REGION Network 10
   RUNG wire#powerrail
      { S7_Templates := "SrcType := Real"; S7_GenerateENO := "TRUE" } Sub(in1 := "DB122".Static_0, in2 := "DB122".Static_24, out => "DB122".Static_18)
      wire#w1
      Coil( "Tag_6" )
   END_RUNG
   RUNG wire#powerrail
      { S7_Templates := "SrcType := Real"; S7_GenerateENO := "TRUE" } Sub(in1 := "DB122".Static_1, in2 := "DB122".Static_24, out => "DB122".Static_19)
   END_RUNG wire#w1
   RUNG wire#powerrail
      { S7_Templates := "SrcType := Real"; S7_GenerateENO := "TRUE" } Sub(in1 := "DB122".Static_2, in2 := "DB122".Static_24, out => "DB122".Static_20)
   END_RUNG wire#w1
   RUNG wire#powerrail
      { S7_Templates := "SrcType := Real"; S7_GenerateENO := "TRUE" } Sub(in1 := "DB122".Static_3, in2 := "DB122".Static_24, out => "DB122".Static_21)
   END_RUNG wire#w1
   RUNG wire#powerrail
      { S7_Templates := "SrcType := Real"; S7_GenerateENO := "TRUE" } Sub(in1 := "DB122".Static_4, in2 := "DB122".Static_24, out => "DB122".Static_22)
   END_RUNG wire#w1
   RUNG wire#powerrail
      { S7_Templates := "SrcType := Real"; S7_GenerateENO := "TRUE" } Sub(in1 := "DB122".Static_5, in2 := "DB122".Static_24, out => "DB122".Static_23)
   END_RUNG wire#w1
   // the same network as SCL:
   // ENO of a box is taken as its EN; it also drops when the box reports an error
   "DB122".Static_18 := "DB122".Static_0 - "DB122".Static_24;
   "DB122".Static_19 := "DB122".Static_1 - "DB122".Static_24;
   "DB122".Static_20 := "DB122".Static_2 - "DB122".Static_24;
   "DB122".Static_21 := "DB122".Static_3 - "DB122".Static_24;
   "DB122".Static_22 := "DB122".Static_4 - "DB122".Static_24;
   "DB122".Static_23 := "DB122".Static_5 - "DB122".Static_24;
   "Tag_6" := TRUE OR TRUE OR TRUE OR TRUE OR TRUE OR TRUE;
END_REGION

REGION Network 11 (STL)
         A     "MC003_EV";
         A(;
         A(;
         L     "DB121".Static_62;
         L     1;
         ==R;
         );
         A(;
         L     "DB52".Static_13;
         L     "DB122".Static_18;
         >=R;
         );
         O;
         A(;
         L     "DB121".Static_62;
         L     2;
         ==R;
         );
         A(;
         L     "DB52".Static_13;
         L     "DB122".Static_19;
         >=R;
         );
         O;
         A(;
         L     "DB121".Static_62;
         L     3;
         ==R;
         );
         A(;
         L     "DB52".Static_13;
         L     "DB122".Static_20;
         >=R;
         );
         O;
         A(;
         L     "DB121".Static_62;
         L     4;
         ==R;
         );
         A(;
         L     "DB52".Static_13;
         L     "DB122".Static_21;
         >=R;
         );
         O;
         A(;
         L     "DB121".Static_62;
         L     5;
         ==R;
         );
         A(;
         L     "DB52".Static_13;
         L     "DB122".Static_22;
         >=R;
         );
         O;
         A(;
         L     "DB121".Static_62;
         L     6;
         ==R;
         );
         A(;
         L     "DB52".Static_13;
         L     "DB122".Static_23;
         >=R;
         );
         );
         L     S5T#30S;
         SF    "Tag_13";
         NOP   0;
         NOP   0;
         NOP   0;
         A     "Tag_13";
         =     #Temp_0;
END_REGION

REGION Network 12
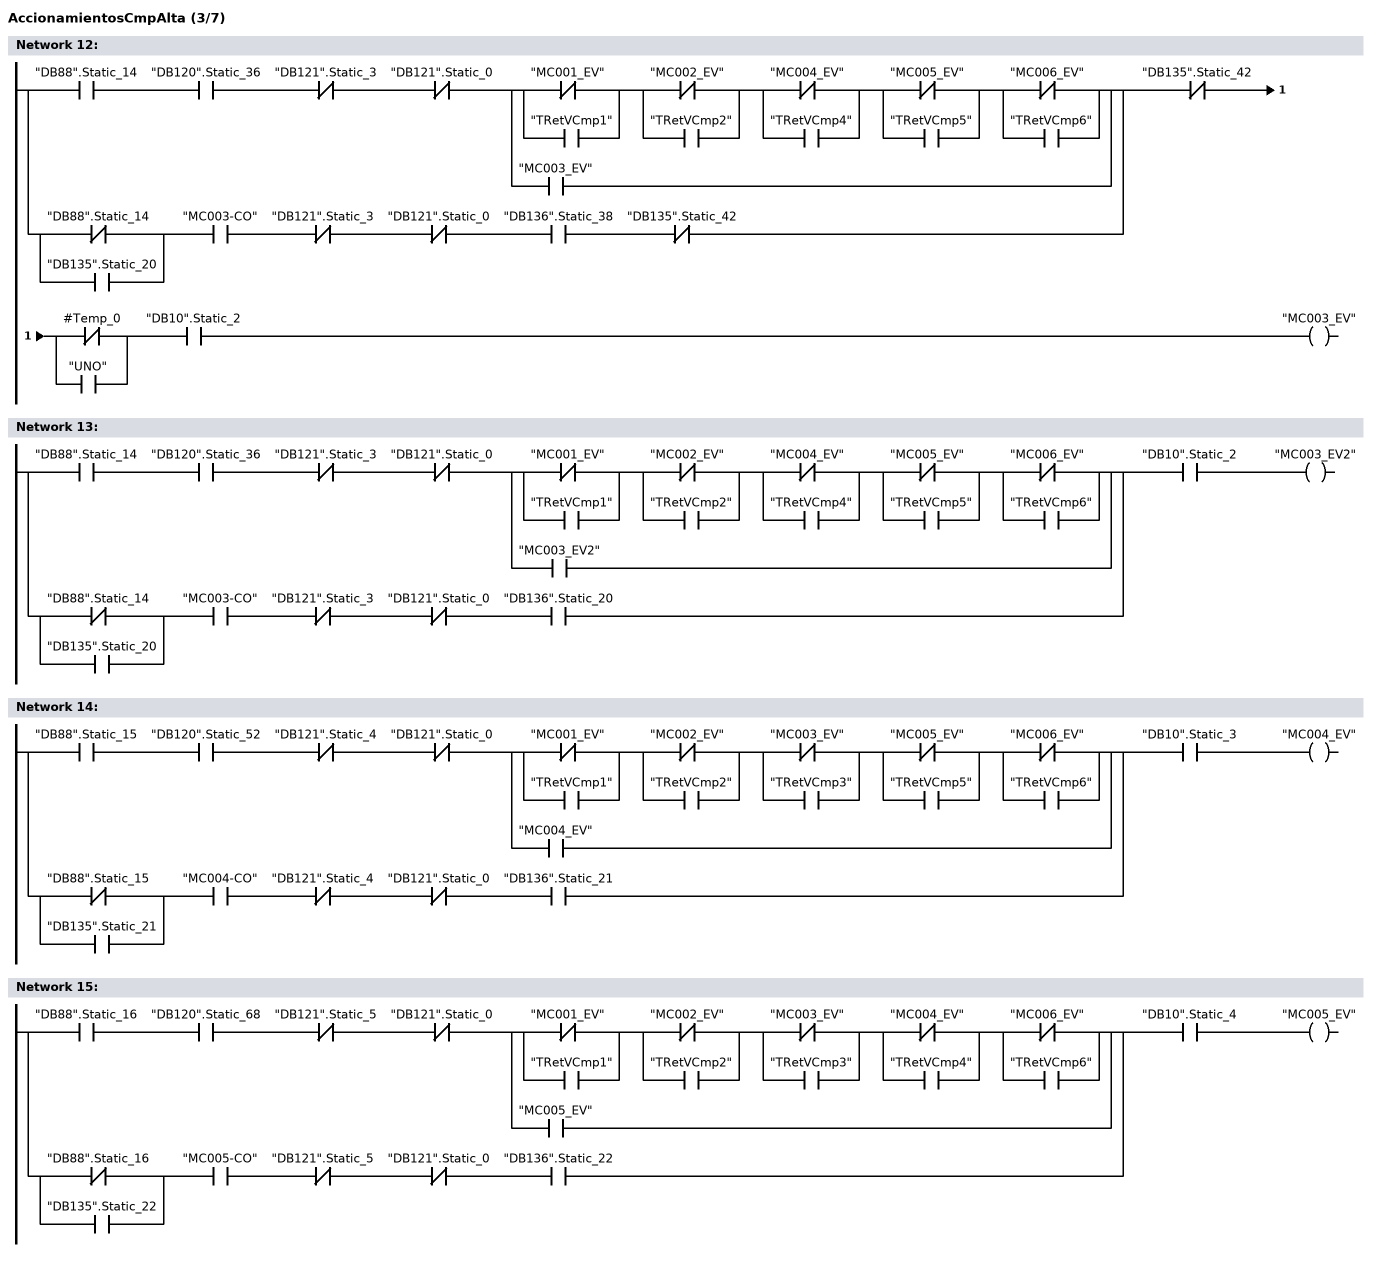
   "MC003_EV" := (("DB88".Static_14 AND "DB120".Static_36 AND NOT "DB121".Static_3 AND NOT "DB121".Static_0 AND (((NOT "MC001_EV" OR "TRetVCmp1") AND (NOT "MC002_EV" OR "TRetVCmp2") AND (NOT "MC004_EV" OR "TRetVCmp4") AND (NOT "MC005_EV" OR "TRetVCmp5") AND (NOT "MC006_EV" OR "TRetVCmp6")) OR "MC003_EV")) OR ((NOT "DB88".Static_14 OR "DB135".Static_20) AND "MC003-CO" AND NOT "DB121".Static_3 AND NOT "DB121".Static_0 AND "DB136".Static_38 AND NOT "DB135".Static_42)) AND NOT "DB135".Static_42 AND (NOT #Temp_0 OR "UNO") AND "DB10".Static_2;
END_REGION

REGION Network 13
   "MC003_EV2" := (("DB88".Static_14 AND "DB120".Static_36 AND NOT "DB121".Static_3 AND NOT "DB121".Static_0 AND (((NOT "MC001_EV" OR "TRetVCmp1") AND (NOT "MC002_EV" OR "TRetVCmp2") AND (NOT "MC004_EV" OR "TRetVCmp4") AND (NOT "MC005_EV" OR "TRetVCmp5") AND (NOT "MC006_EV" OR "TRetVCmp6")) OR "MC003_EV2")) OR ((NOT "DB88".Static_14 OR "DB135".Static_20) AND "MC003-CO" AND NOT "DB121".Static_3 AND NOT "DB121".Static_0 AND "DB136".Static_20)) AND "DB10".Static_2;
END_REGION

REGION Network 14
   "MC004_EV" := (("DB88".Static_15 AND "DB120".Static_52 AND NOT "DB121".Static_4 AND NOT "DB121".Static_0 AND (((NOT "MC001_EV" OR "TRetVCmp1") AND (NOT "MC002_EV" OR "TRetVCmp2") AND (NOT "MC003_EV" OR "TRetVCmp3") AND (NOT "MC005_EV" OR "TRetVCmp5") AND (NOT "MC006_EV" OR "TRetVCmp6")) OR "MC004_EV")) OR ((NOT "DB88".Static_15 OR "DB135".Static_21) AND "MC004-CO" AND NOT "DB121".Static_4 AND NOT "DB121".Static_0 AND "DB136".Static_21)) AND "DB10".Static_3;
END_REGION

REGION Network 15
   "MC005_EV" := (("DB88".Static_16 AND "DB120".Static_68 AND NOT "DB121".Static_5 AND NOT "DB121".Static_0 AND (((NOT "MC001_EV" OR "TRetVCmp1") AND (NOT "MC002_EV" OR "TRetVCmp2") AND (NOT "MC003_EV" OR "TRetVCmp3") AND (NOT "MC004_EV" OR "TRetVCmp4") AND (NOT "MC006_EV" OR "TRetVCmp6")) OR "MC005_EV")) OR ((NOT "DB88".Static_16 OR "DB135".Static_22) AND "MC005-CO" AND NOT "DB121".Static_5 AND NOT "DB121".Static_0 AND "DB136".Static_22)) AND "DB10".Static_4;
END_REGION

REGION Network 16
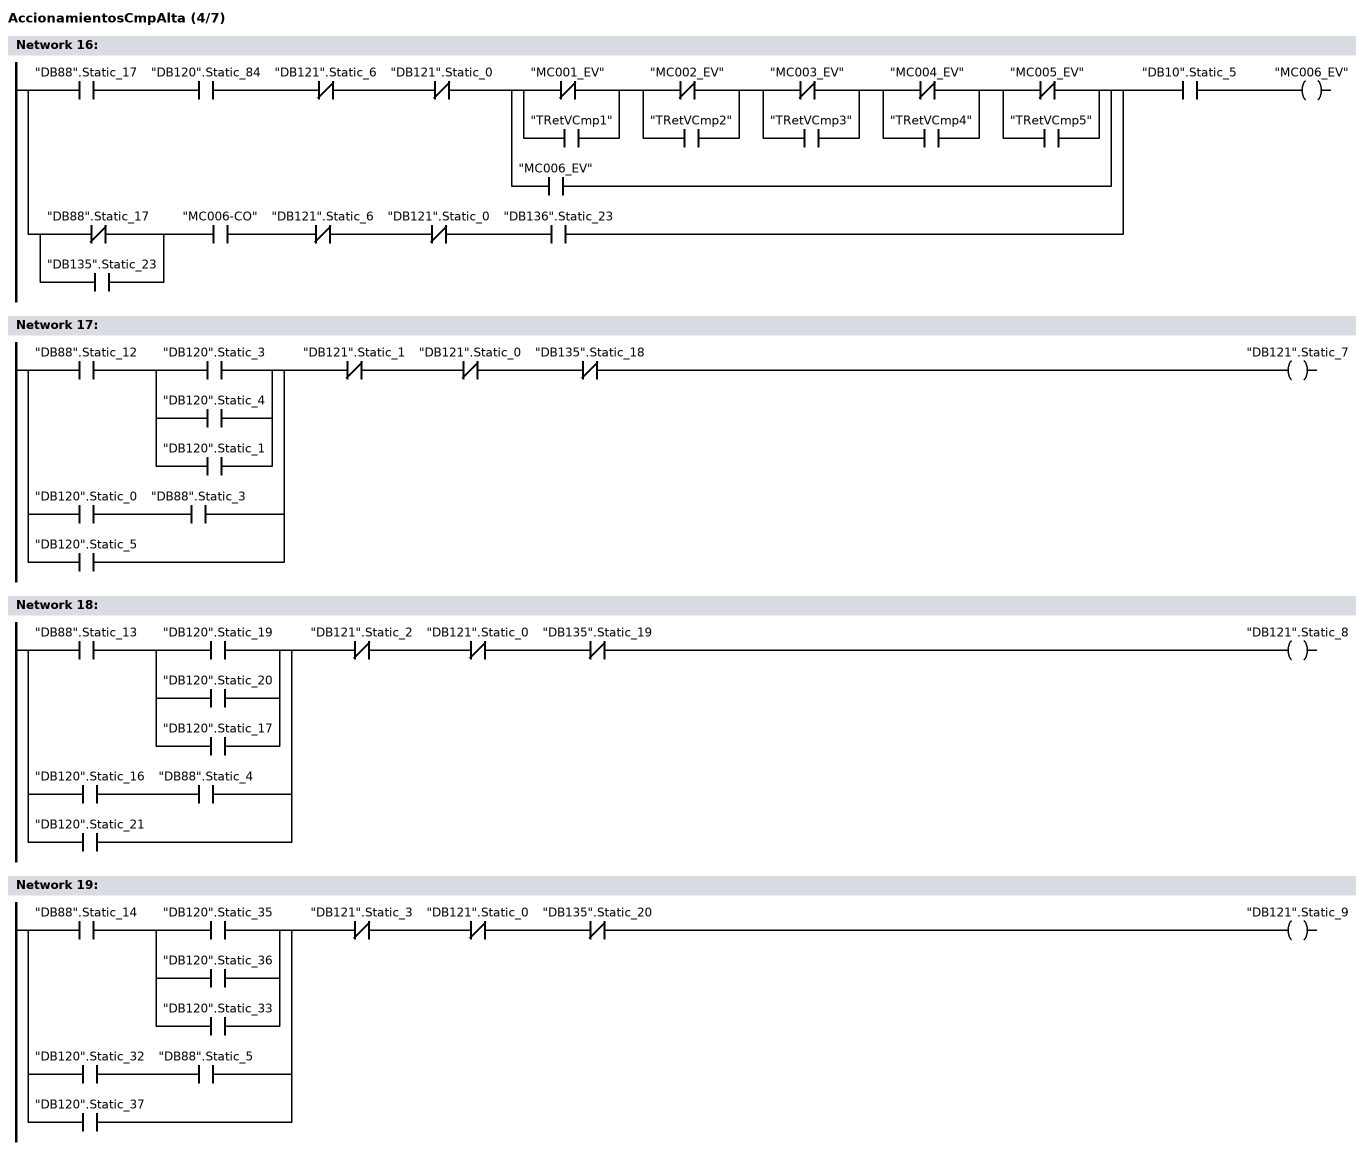
   "MC006_EV" := (("DB88".Static_17 AND "DB120".Static_84 AND NOT "DB121".Static_6 AND NOT "DB121".Static_0 AND (((NOT "MC001_EV" OR "TRetVCmp1") AND (NOT "MC002_EV" OR "TRetVCmp2") AND (NOT "MC003_EV" OR "TRetVCmp3") AND (NOT "MC004_EV" OR "TRetVCmp4") AND (NOT "MC005_EV" OR "TRetVCmp5")) OR "MC006_EV")) OR ((NOT "DB88".Static_17 OR "DB135".Static_23) AND "MC006-CO" AND NOT "DB121".Static_6 AND NOT "DB121".Static_0 AND "DB136".Static_23)) AND "DB10".Static_5;
END_REGION

REGION Network 17
   "DB121".Static_7 := (("DB88".Static_12 AND ("DB120".Static_3 OR "DB120".Static_4 OR "DB120".Static_1)) OR ("DB120".Static_0 AND "DB88".Static_3) OR "DB120".Static_5) AND NOT "DB121".Static_1 AND NOT "DB121".Static_0 AND NOT "DB135".Static_18;
END_REGION

REGION Network 18
   "DB121".Static_8 := (("DB88".Static_13 AND ("DB120".Static_19 OR "DB120".Static_20 OR "DB120".Static_17)) OR ("DB120".Static_16 AND "DB88".Static_4) OR "DB120".Static_21) AND NOT "DB121".Static_2 AND NOT "DB121".Static_0 AND NOT "DB135".Static_19;
END_REGION

REGION Network 19
   "DB121".Static_9 := (("DB88".Static_14 AND ("DB120".Static_35 OR "DB120".Static_36 OR "DB120".Static_33)) OR ("DB120".Static_32 AND "DB88".Static_5) OR "DB120".Static_37) AND NOT "DB121".Static_3 AND NOT "DB121".Static_0 AND NOT "DB135".Static_20;
END_REGION

REGION Network 20
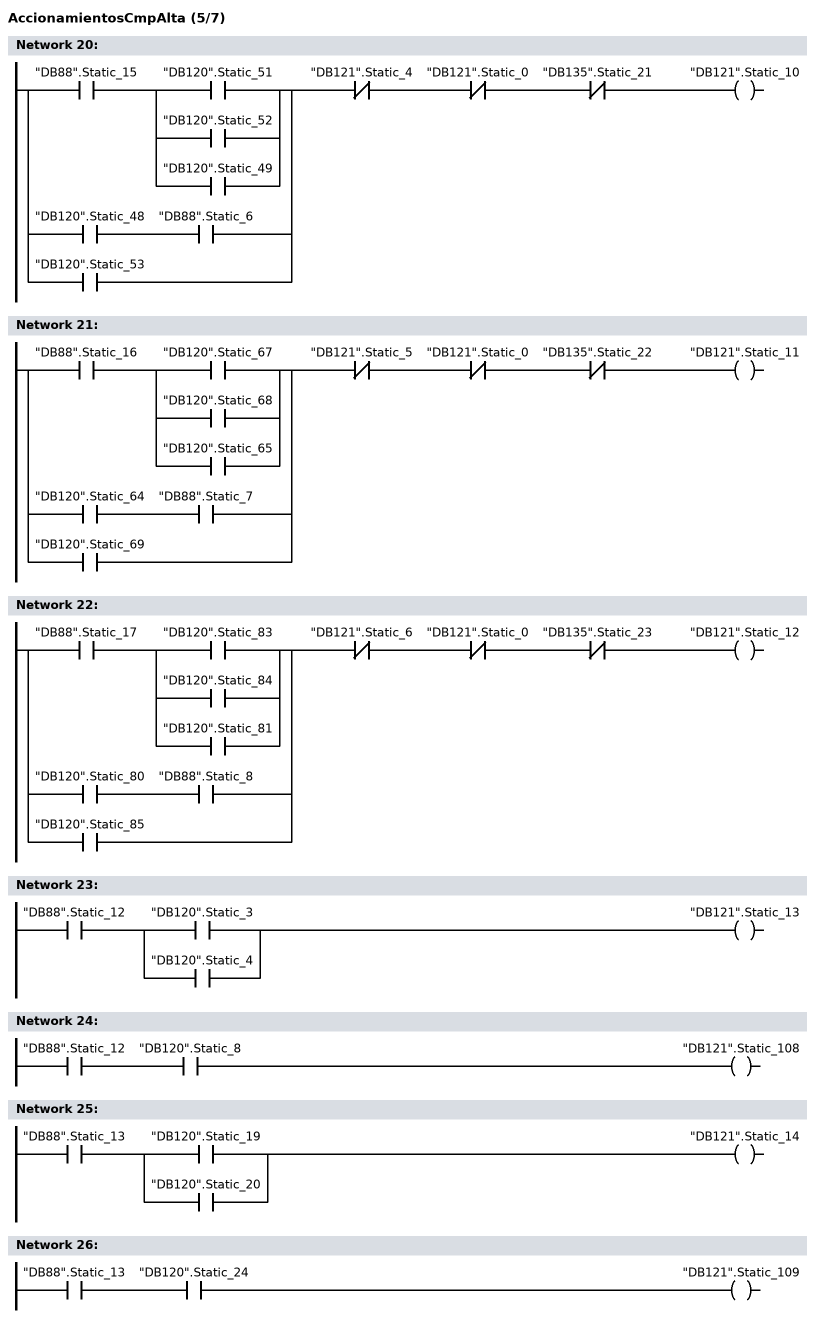
   "DB121".Static_10 := (("DB88".Static_15 AND ("DB120".Static_51 OR "DB120".Static_52 OR "DB120".Static_49)) OR ("DB120".Static_48 AND "DB88".Static_6) OR "DB120".Static_53) AND NOT "DB121".Static_4 AND NOT "DB121".Static_0 AND NOT "DB135".Static_21;
END_REGION

REGION Network 21
   "DB121".Static_11 := (("DB88".Static_16 AND ("DB120".Static_67 OR "DB120".Static_68 OR "DB120".Static_65)) OR ("DB120".Static_64 AND "DB88".Static_7) OR "DB120".Static_69) AND NOT "DB121".Static_5 AND NOT "DB121".Static_0 AND NOT "DB135".Static_22;
END_REGION

REGION Network 22
   "DB121".Static_12 := (("DB88".Static_17 AND ("DB120".Static_83 OR "DB120".Static_84 OR "DB120".Static_81)) OR ("DB120".Static_80 AND "DB88".Static_8) OR "DB120".Static_85) AND NOT "DB121".Static_6 AND NOT "DB121".Static_0 AND NOT "DB135".Static_23;
END_REGION

REGION Network 23
   "DB121".Static_13 := "DB88".Static_12 AND ("DB120".Static_3 OR "DB120".Static_4);
END_REGION

REGION Network 24
   RUNG wire#powerrail
      Contact( "DB88".Static_12 )
      Contact( "DB120".Static_8 )
      Coil( "DB121".Static_108 )
   END_RUNG
   // the same network as SCL:
   "DB121".Static_108 := "DB88".Static_12 AND "DB120".Static_8;
END_REGION

REGION Network 25
   "DB121".Static_14 := "DB88".Static_13 AND ("DB120".Static_19 OR "DB120".Static_20);
END_REGION

REGION Network 26
   RUNG wire#powerrail
      Contact( "DB88".Static_13 )
      Contact( "DB120".Static_24 )
      Coil( "DB121".Static_109 )
   END_RUNG
   // the same network as SCL:
   "DB121".Static_109 := "DB88".Static_13 AND "DB120".Static_24;
END_REGION

REGION Network 27
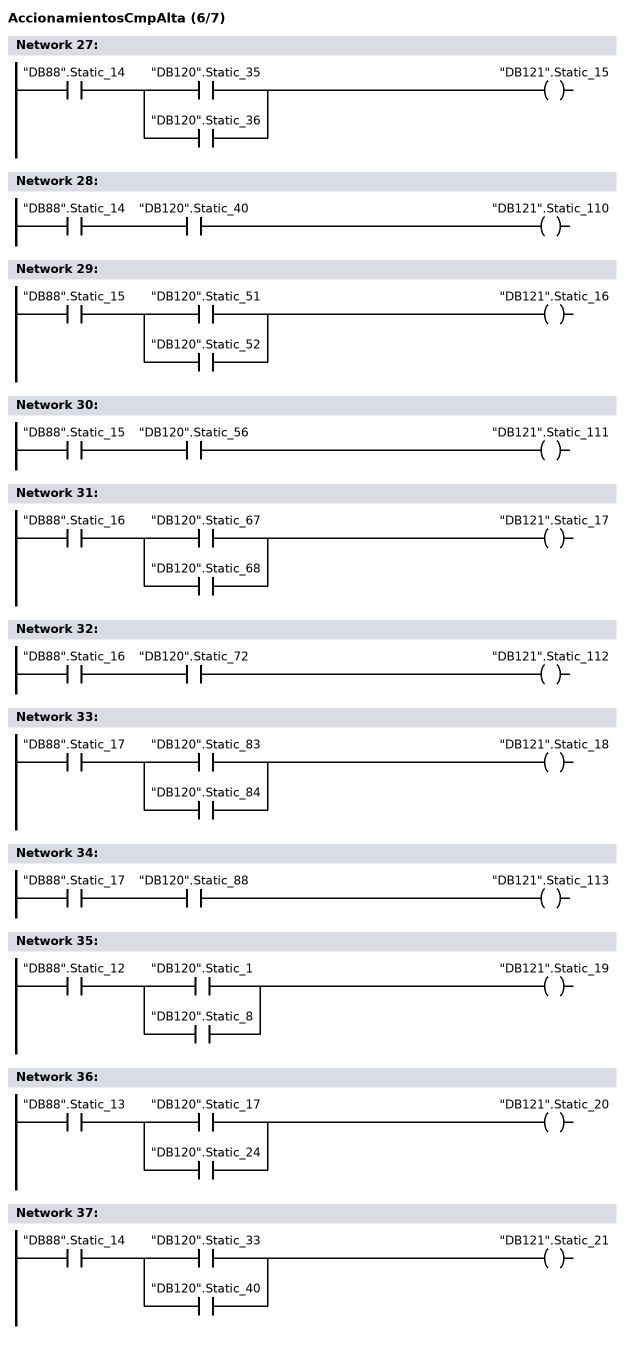
   "DB121".Static_15 := "DB88".Static_14 AND ("DB120".Static_35 OR "DB120".Static_36);
END_REGION

REGION Network 28
   RUNG wire#powerrail
      Contact( "DB88".Static_14 )
      Contact( "DB120".Static_40 )
      Coil( "DB121".Static_110 )
   END_RUNG
   // the same network as SCL:
   "DB121".Static_110 := "DB88".Static_14 AND "DB120".Static_40;
END_REGION

REGION Network 29
   "DB121".Static_16 := "DB88".Static_15 AND ("DB120".Static_51 OR "DB120".Static_52);
END_REGION

REGION Network 30
   RUNG wire#powerrail
      Contact( "DB88".Static_15 )
      Contact( "DB120".Static_56 )
      Coil( "DB121".Static_111 )
   END_RUNG
   // the same network as SCL:
   "DB121".Static_111 := "DB88".Static_15 AND "DB120".Static_56;
END_REGION

REGION Network 31
   "DB121".Static_17 := "DB88".Static_16 AND ("DB120".Static_67 OR "DB120".Static_68);
END_REGION

REGION Network 32
   RUNG wire#powerrail
      Contact( "DB88".Static_16 )
      Contact( "DB120".Static_72 )
      Coil( "DB121".Static_112 )
   END_RUNG
   // the same network as SCL:
   "DB121".Static_112 := "DB88".Static_16 AND "DB120".Static_72;
END_REGION

REGION Network 33
   "DB121".Static_18 := "DB88".Static_17 AND ("DB120".Static_83 OR "DB120".Static_84);
END_REGION

REGION Network 34
   RUNG wire#powerrail
      Contact( "DB88".Static_17 )
      Contact( "DB120".Static_88 )
      Coil( "DB121".Static_113 )
   END_RUNG
   // the same network as SCL:
   "DB121".Static_113 := "DB88".Static_17 AND "DB120".Static_88;
END_REGION

REGION Network 35
   "DB121".Static_19 := "DB88".Static_12 AND ("DB120".Static_1 OR "DB120".Static_8);
END_REGION

REGION Network 36
   "DB121".Static_20 := "DB88".Static_13 AND ("DB120".Static_17 OR "DB120".Static_24);
END_REGION

REGION Network 37
   "DB121".Static_21 := "DB88".Static_14 AND ("DB120".Static_33 OR "DB120".Static_40);
END_REGION

REGION Network 38
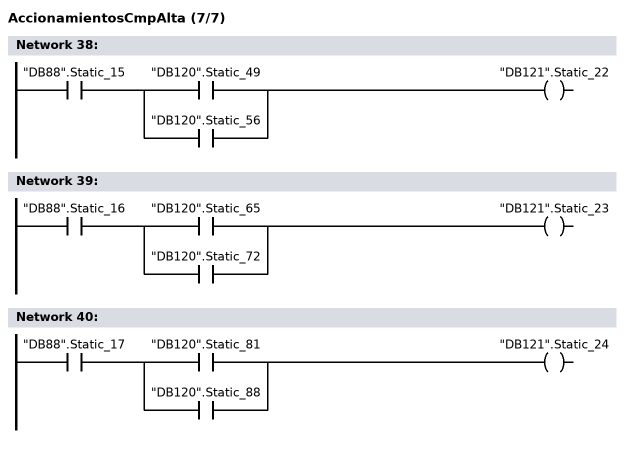
   "DB121".Static_22 := "DB88".Static_15 AND ("DB120".Static_49 OR "DB120".Static_56);
END_REGION

REGION Network 39
   "DB121".Static_23 := "DB88".Static_16 AND ("DB120".Static_65 OR "DB120".Static_72);
END_REGION

REGION Network 40
   "DB121".Static_24 := "DB88".Static_17 AND ("DB120".Static_81 OR "DB120".Static_88);
END_REGION
END_FUNCTION

FUNCTION "PrioridadesReales" : Void   // FC41, LAD
{ S7_Optimized_Access := 'FALSE' }
VERSION : 0.1
BEGIN

REGION Network 1
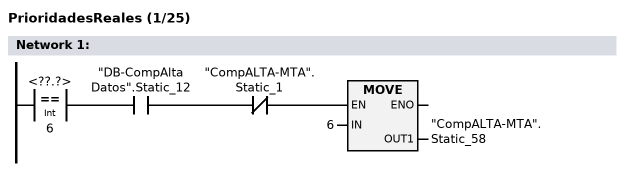
   RUNG wire#powerrail
      { S7_Templates := "SrcType := Int" } EQ_Contact(in1 :=, in2 := 6)
      Contact( "DB-CompAltaDatos".Static_12 )
      I_Contact( "CompALTA-MTA".Static_1 )
      { S7_GenerateENO := "TRUE" } Move(in := 6, out1 => "CompALTA-MTA".Static_58)
   END_RUNG
   // the same network as SCL:
   IF (<??.?> = 6) AND "DB-CompAltaDatos".Static_12 AND NOT "CompALTA-MTA".Static_1 THEN
       "CompALTA-MTA".Static_58 := 6;
   END_IF;
END_REGION

REGION Network 2
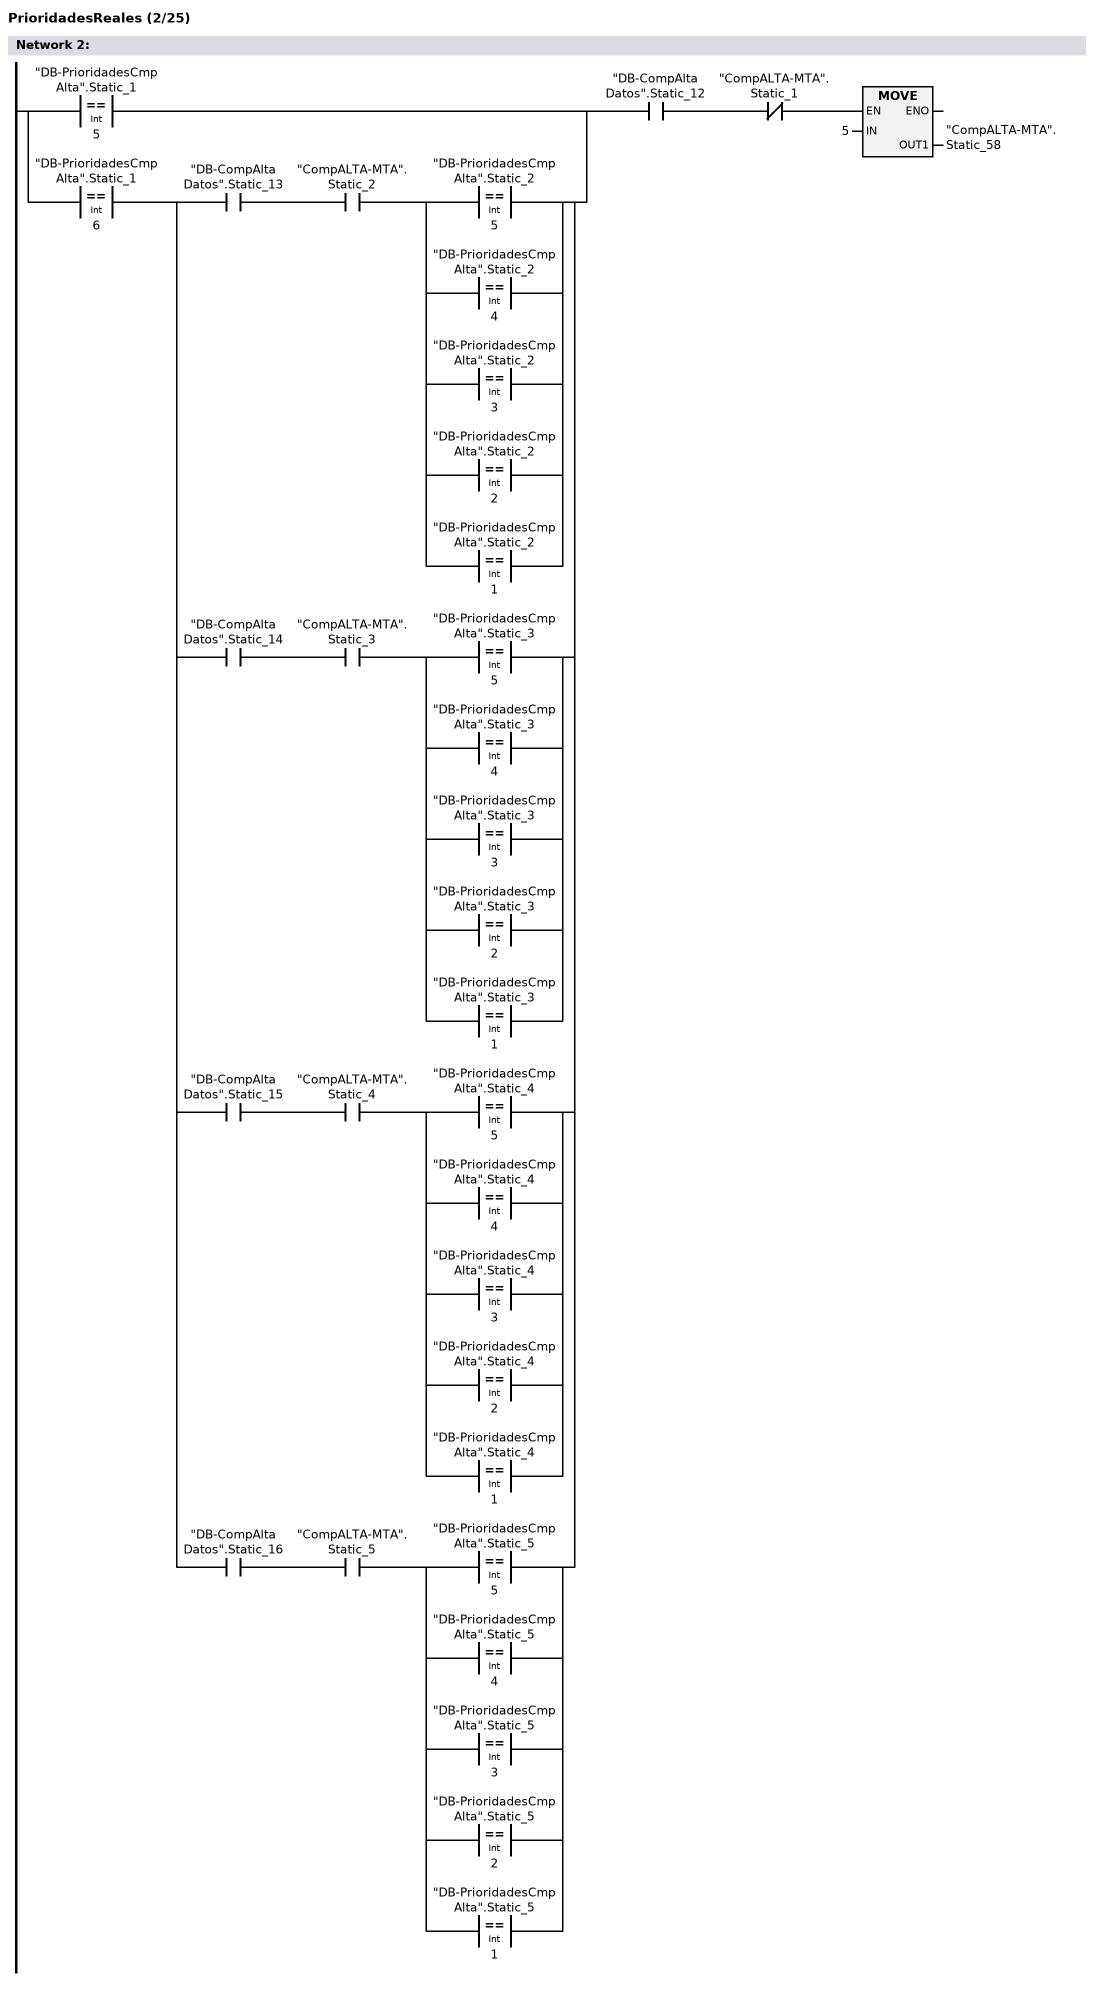
   IF (("DB-PrioridadesCmpAlta".Static_1 = 5) OR (("DB-PrioridadesCmpAlta".Static_1 = 6) AND (("DB-CompAltaDatos".Static_13 AND "CompALTA-MTA".Static_2 AND (("DB-PrioridadesCmpAlta".Static_2 = 5) OR ("DB-PrioridadesCmpAlta".Static_2 = 4) OR ("DB-PrioridadesCmpAlta".Static_2 = 3) OR ("DB-PrioridadesCmpAlta".Static_2 = 2) OR ("DB-PrioridadesCmpAlta".Static_2 = 1))) OR ("DB-CompAltaDatos".Static_14 AND "CompALTA-MTA".Static_3 AND (("DB-PrioridadesCmpAlta".Static_3 = 5) OR ("DB-PrioridadesCmpAlta".Static_3 = 4) OR ("DB-PrioridadesCmpAlta".Static_3 = 3) OR ("DB-PrioridadesCmpAlta".Static_3 = 2) OR ("DB-PrioridadesCmpAlta".Static_3 = 1))) OR ("DB-CompAltaDatos".Static_15 AND "CompALTA-MTA".Static_4 AND (("DB-PrioridadesCmpAlta".Static_4 = 5) OR ("DB-PrioridadesCmpAlta".Static_4 = 4) OR ("DB-PrioridadesCmpAlta".Static_4 = 3) OR ("DB-PrioridadesCmpAlta".Static_4 = 2) OR ("DB-PrioridadesCmpAlta".Static_4 = 1))) OR ("DB-CompAltaDatos".Static_16 AND "CompALTA-MTA".Static_5 AND (("DB-PrioridadesCmpAlta".Static_5 = 5) OR ("DB-PrioridadesCmpAlta".Static_5 = 4) OR ("DB-PrioridadesCmpAlta".Static_5 = 3) OR ("DB-PrioridadesCmpAlta".Static_5 = 2) OR ("DB-PrioridadesCmpAlta".Static_5 = 1)))))) AND "DB-CompAltaDatos".Static_12 AND NOT "CompALTA-MTA".Static_1 THEN
       "CompALTA-MTA".Static_58 := 5;
   END_IF;
END_REGION

REGION Network 3
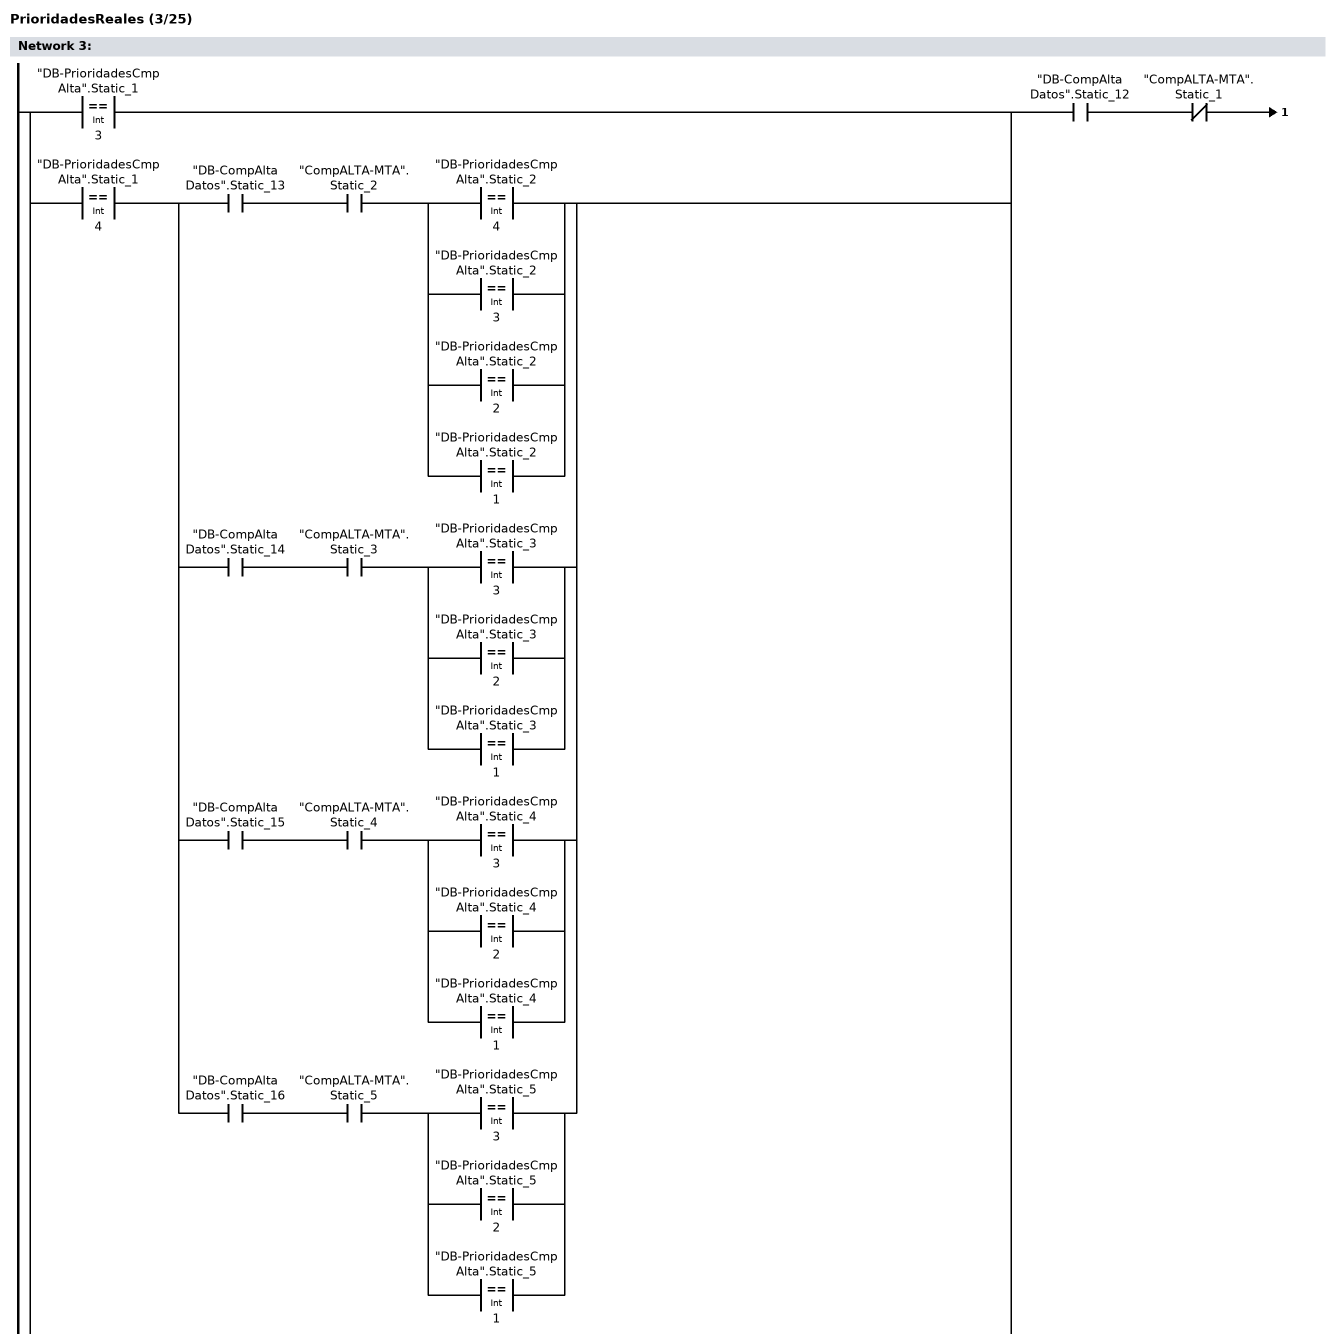
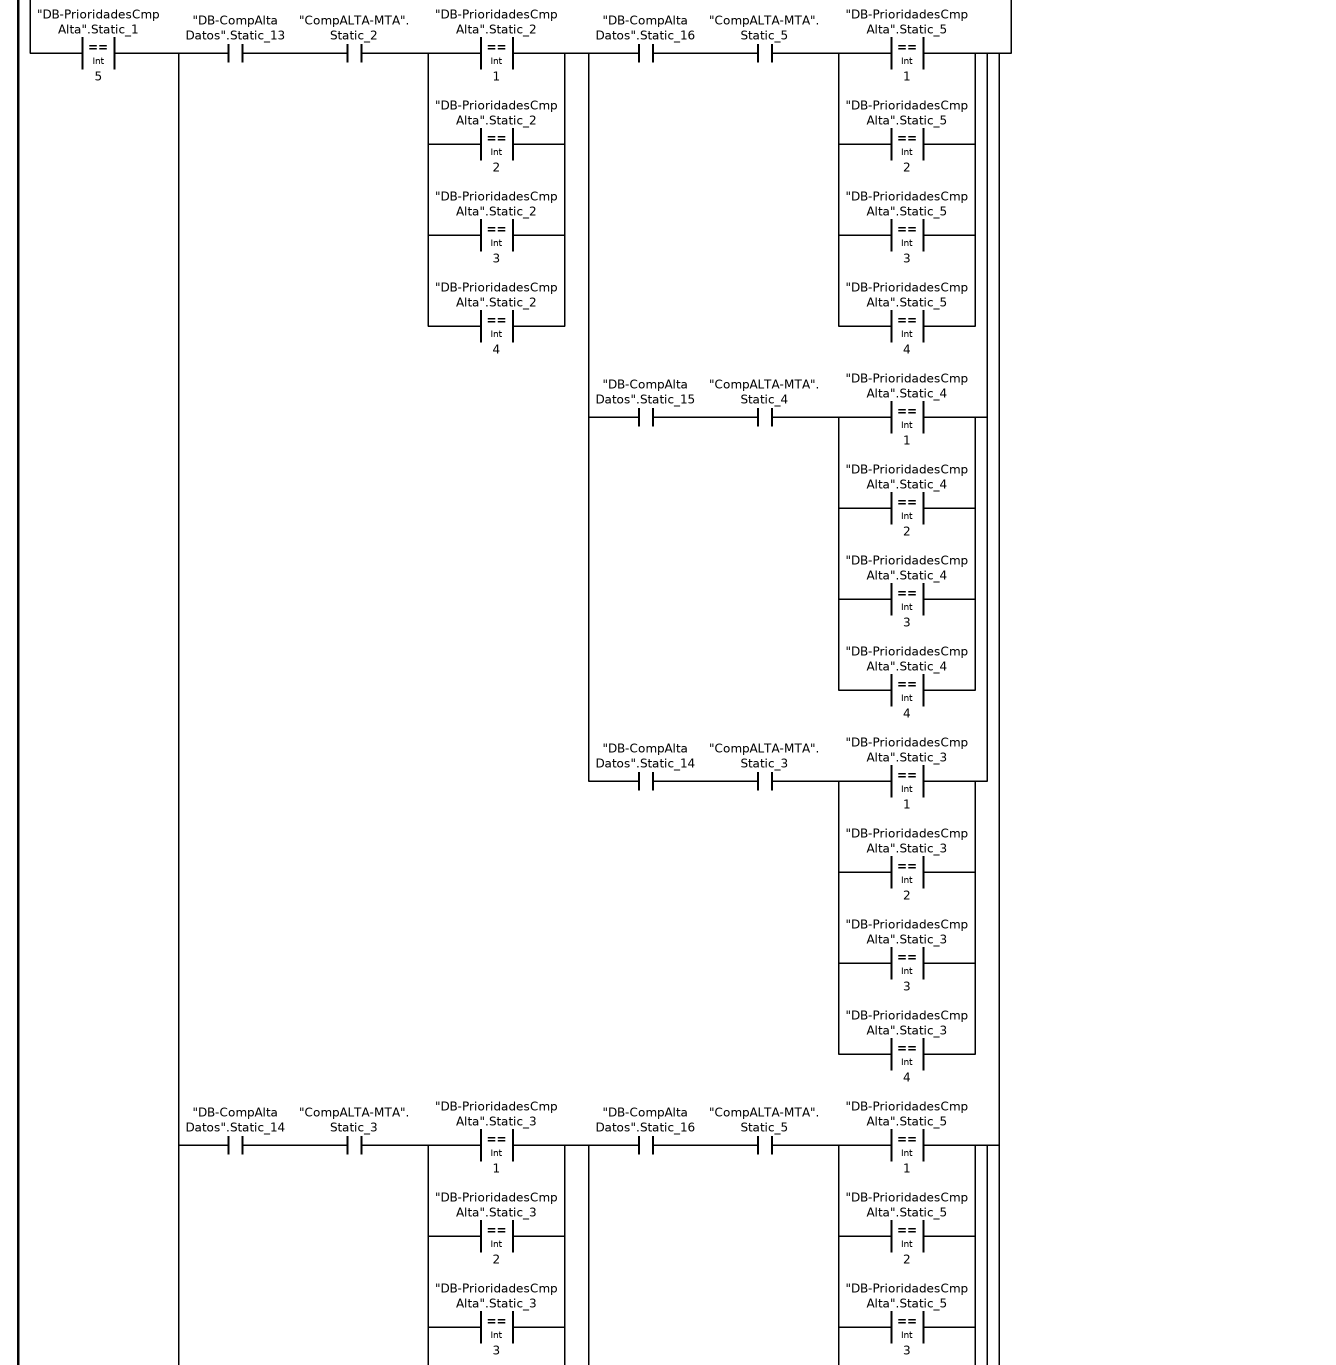
